
     ELSIF (#statStatus = #STATUS_COMMAND_ABORTED) AND (#statCommandAborted = FALSE) THEN // Commanded functionality has been aborted by another command
       #statDone := FALSE;
       #statBusy := FALSE;
       #statCommandAborted := TRUE;
       #statError := FALSE;
       #diagnostics.stateNumber := #statFBState;
       #diagnostics.status := #statStatus;
       #diagnostics.subfunctionStatus := #statSubfunctionStatus;
       #statFBState := #FB_STATE_NO_PROCESSING; // Switch state machine to "no processing"

       // Reset pointer
       #lineBuffer.pointers.addPointer := 0;
       #lineBuffer.pointers.addPointerRestarted := FALSE;
       #lineBuffer.pointers.bufferLocked := FALSE;
       IF #lineBuffer.info.fileState <> "LKINLANG_FILE_STATE_RUNNING"
         AND #lineBuffer.info.fileState <> "LKINLANG_FILE_STATE_RUNNING_LOADING" THEN
         #lineBuffer.pointers.ignoreAddPointer := TRUE;
       END_IF;

       // Set file state
       #lineBuffer.info.fileState := "LKINLANG_FILE_STATE_STOPPED";


     ELSIF (#statCommandAborted = TRUE) AND (#tempStop = FALSE) THEN
       #statDone := FALSE;
       #statBusy := FALSE;
       #statCommandAborted := FALSE;
       #statError := FALSE;
       #statStatus := #STATUS_NO_CALL;

       // Reset file state
       #lineBuffer.info.fileState := "LKINLANG_FILE_STATE_IDLE";

     ELSIF (#tempExecuteCardToPlc = FALSE) AND (#tempExecutePlcToCard = FALSE) AND ((#statDone = TRUE) OR (#statError = TRUE)) THEN
       #statDone := FALSE;
       #statBusy := FALSE;
       #statCommandAborted := FALSE;
       #statError := FALSE;
       #statStatus := #STATUS_NO_CALL;

       IF #lineBuffer.info.fileState = "LKINLANG_FILE_STATE_STOPPED" THEN
         // Reset file state
         #lineBuffer.info.fileState := "LKINLANG_FILE_STATE_IDLE";
       END_IF;
     END_IF;


     // Write static values to outputs
     #done := #statDone;
     #busy := #statBusy;
     #dataTransferStopped := #statCommandAborted;
     #error := #statError;
     #status := #statStatus;

   END_REGION OUTPUTS

   //--------------------------------------------------------------------
   // End of Block LKinLang_FileHandler
   //--------------------------------------------------------------------
END_FUNCTION_BLOCK

FUNCTION_BLOCK "LKinLang_ProgramLineDisplay"   // FB35452, SCL
TITLE = LKinLang_ProgramLineDisplay
{ S7_Optimized_Access := 'TRUE' }
AUTHOR : tech.team.motioncontrol@siemens.com
FAMILY : LKinLang
VERSION : 1.0
// This FB shows the current parsed, buffered and active line
   VAR_INPUT
      enable : Bool;   // TRUE: Enable functionality of FB
      activeCmdNo : DInt;   // Currently active command number (FB MovePath output)
      movePathStatus : Word;   // Current status output of FB MovePath
   END_VAR
   VAR_OUTPUT
      valid : Bool;   // TRUE: Valid set of output values available at the FB
      busy : Bool;   // TRUE: FB is not finished and new output values can be expected
      error : Bool;   // TRUE: An error occurred during the execution of the FB
      status : Word := 16#7000;   // 16#0000 - 16#7FFF: Status of the FB, 16#8000 - 16#FFFF: Error identification
      parsedLineNo : UDInt;   // Last parsed line number
      parsedLine : String;   // Last parsed line
      bufferedLineNo : UDInt;   // Last buffered line number (internal storage of FB MovePath)
      bufferedLine : String;   // Last buffered line (internal storage of FB MovePath)
      activeLineNo : UDInt;   // Currently active line number
      activeLine : String;   // Currently active line
   END_VAR
   VAR_IN_OUT
      lineBuffer : "LKinLang_typeLineBuffer";   // LineBuffer connection
      pathData : "LKinCtrl_typePathData_advanced";   // PathData connection
   END_VAR
   VAR
      statEnableOld : Bool;   // Old value of 'enable' input for edge detection
      statValid : Bool;   // Static value for output 'valid'
      statBusy : Bool;   // Static value for output 'busy'
      statError : Bool;   // Static value for output 'error'
      statStatus : Word := 16#7000;   // Static value for output 'status'
      statParsedLine : String;   // Static value for output 'parsedLine'
      statParsedLineNo : UDInt;   // Static value for output 'parsedLineNo'
      statBufferedLine : String;   // Static value for output 'bufferedLine'
      statBufferedLineNo : UDInt;   // Static value for output 'bufferedLineNo'
      statActiveLine : String;   // Static value for output 'activeLine'
      statActiveLineNo : UDInt;   // Static value for output 'activeLineNo'
      statErrorUserCleared : Bool;   // Error occurred that can only be solved by user; rising edge at enable input necessary
      statErrorAutoCleared : Bool;   // Error occurred that can be acknowledged by FB
      statFBState : DInt := 0;   // State in the state machine of the FB
      statDisablingCompleted : Bool;   // TRUE: Disabling has been completed
      statAddPointerPathOld : DInt;   // Last value of PathData add pointer
      statRetPointerPathOld : DInt;   // Last value of PathData retrieve pointer
      statActiveCmdNoOld : DInt;   // Last value of active command number
      statRetPointerLineOld : DInt;   // Last value of LineBuffer retrieve pointer
      statBufferIndex : DInt;   // Counter for internal buffer
      statFirstBufferEntry : DInt;   // Static storage for first entry in internal buffer
      statFirstActiveBufferEntry : DInt;   // Static storage for first active entry in internal buffer
      statParsingDone : Bool;   // TRUE: FB Parser is done
      statBufferingDone : Bool;   // TRUE: FB MovePath has copied all commands from PathData
      statMovePathDone : Bool;   // TRUE: FB MovePath has executed all commands from PathData
      statPathDataLines : Array[1.."LKINCTRL_NO_OF_PATHDATA_ELEMENTS_ADVANCED"] of String["LKINLANG_LENGTH_OF_ASCII_LINE_STRING"];   // Stores the corresponding lines from PathData
      statPathDataLineNo : Array[1.."LKINCTRL_NO_OF_PATHDATA_ELEMENTS_ADVANCED"] of UDInt;   // Stores the corresponding line numbers from PathData
      statInternalLines : Array[0..#LAST_INDEX_INTERNAL] of String["LKINLANG_LENGTH_OF_ASCII_LINE_STRING"];   // Stores the corresponding lines from FB MovePath internal buffer
      statInternalLineNo : Array[0..#LAST_INDEX_INTERNAL] of UDInt;   // Stores the corresponding line numbers from FB MovePath internal buffer
   END_VAR
   VAR_TEMP
      tempEnable : Bool;   // Temporary value for input 'enable'
      tempAddPointerPath : DInt;   // Temporary value for input 'PathData.pointers.addPointer'
      tempRetPointerPath : DInt;   // Temporary value for input 'PathData.pointers.retrievePointer'
      tempAddPointerLine : DInt;   // Temporary value for input 'LineBuffer.pointers.addPointer'
      tempRetPointerLine : DInt;   // Temporary value for input 'LineBuffer.pointers.retrievePointer'
      tempActiveCmdNo : DInt;   // Temporary value for input 'activeCmdNo'
      tempMovePathStatus : DWord;   // Temporary value for input 'movePathStatus'
      tempIndex : DInt;   // Temporary counter
   END_VAR
   VAR CONSTANT
      FB_STATE_NO_PROCESSING : DInt := 0;   // FB state: No processing
      FB_STATE_PROCESSING : DInt := 50;   // FB state: Processing
      FB_STATE_DISABLING : DInt := 90;   // FB state: Disabling
      STATUS_NO_CALL : Word := 16#7000;   // No job being currently processed
      STATUS_FIRST_CALL : Word := 16#7001;   // First call after incoming new job (rising edge 'enable')
      STATUS_SUBSEQUENT_CALL : Word := 16#7002;   // Subsequent call during active processing without further details
      ERR_UNDEFINED_STATE : Word := 16#8600;   // Error due to an undefined state in state machine
      LAST_INDEX_INTERNAL : DInt := 19;   // Last index of internal array
   END_VAR
BEGIN
   //=============================================================================
   // SIEMENS AG
   // (c)Copyright 2020
   //-----------------------------------------------------------------------------
   // Library:       LKinLang
   // Tested with:   S7-1517T-3 PN/DP
   // Engineering:   TIA Portal V16
   // Restrictions:  -
   // Requirements:  -
   // Functionality: This FB shows the current parsed, buffered and active line
   //-----------------------------------------------------------------------------
   // Change log table:
   // Version      Date        Expert in charge    Changes applied
   // 01.00.00     03.12.2020  FR                  First created version
   //=============================================================================

   // Work with temporary value / create process image
   #tempEnable := #enable;
   #tempAddPointerPath := #pathData.pointers.addPointer;
   #tempRetPointerPath := #pathData.pointers.retrievePointer;
   #tempAddPointerLine := #lineBuffer.pointers.addPointer;
   #tempRetPointerLine := #lineBuffer.pointers.retrievePointer;
   #tempActiveCmdNo := #activeCmdNo;
   #tempMovePathStatus := #movePathStatus;

   REGION ENABLING/DISABLING
       IF (#tempEnable = TRUE) AND (#statStatus = #STATUS_NO_CALL) THEN // Enable FB
           // First call; initialize FB
           #statValid := TRUE;
           #statBusy := TRUE;
           #statError := FALSE;
           #statErrorUserCleared := FALSE;
           #statErrorAutoCleared := FALSE;
           #statStatus := #STATUS_FIRST_CALL;

           #statFBState := #FB_STATE_PROCESSING; // State machine - start functionality

           // Reset of variables, diagnostics, etc.
           #statDisablingCompleted := FALSE;

           // Reset "old" variables
           #statAddPointerPathOld := 0;
           #statRetPointerPathOld := 0;
           #statActiveCmdNoOld := 0;
           #statRetPointerLineOld := 0;

           // Reset counter / index
           #statBufferIndex := 0;
           #statFirstBufferEntry := 0;
           #statFirstActiveBufferEntry := 0;

           // Reset status bits
           #statParsingDone := FALSE;
           #statBufferingDone := FALSE;

           // Reset arrays
           FOR #tempIndex := 0 TO #LAST_INDEX_INTERNAL DO
               #statInternalLines[#tempIndex] := '';
               #statInternalLineNo[#tempIndex] := 0;
           END_FOR;
           FOR #tempIndex := 1 TO "LKINCTRL_NO_OF_PATHDATA_ELEMENTS_ADVANCED" DO
               #statPathDataLines[#tempIndex] := '';
               #statPathDataLineNo[#tempIndex] := 0;
           END_FOR;

       ELSIF (#tempEnable = FALSE) AND (#statEnableOld = TRUE) THEN // Disable FB 
           #statFBState := #FB_STATE_DISABLING;

       ELSIF (#statStatus = #STATUS_FIRST_CALL) THEN // Set status identifier of subsequent call
           #statStatus := #STATUS_SUBSEQUENT_CALL;
       END_IF;

       // Edge detection 'enable' input
       #statEnableOld := #tempEnable;
   END_REGION ENABLING/DISABLING

   IF (#statStatus = #STATUS_NO_CALL) THEN // Nothing to do -> End here to reduce "system load"
       RETURN;
   END_IF;

   REGION STATE_MACHINE
       CASE #statFBState OF // State machine of FB
           #FB_STATE_NO_PROCESSING: // No processing active (Note: this state must always be present and left empty)
               ;

           #FB_STATE_PROCESSING: // Processing active
               // -----------------------------------------------------------------
               // If a new pathData command was added then store the corresponding
               // lineBuffer entry in the internal pathData buffer
               // 
               // Also check if parsing has finished
               // -----------------------------------------------------------------
               REGION STORE_LINES_INTERNAL
                   // Calculate index
                   IF #tempRetPointerLine > 0 THEN
                       // regular 
                       #tempIndex := #tempRetPointerLine;
                       #statParsingDone := FALSE;
                   ELSIF #tempRetPointerLine = 0 AND #statRetPointerLineOld <> 0 THEN
                       // Parser finished --> retrieve pointer is reset instantly --> Use old value
                       #tempIndex := #statRetPointerLineOld;
                       #statParsingDone := TRUE;
                   ELSE
                       #tempIndex := 0;
                   END_IF;

                   // Check if new pathData command was added
                   IF #tempAddPointerPath <> #statAddPointerPathOld AND #tempAddPointerPath > 0 AND #tempIndex <> 0 THEN
                       // Store the corresponding line in path data line buffer
                       #statPathDataLines[#tempAddPointerPath] := #lineBuffer.lines[#tempIndex].content;
                       #statPathDataLineNo[#tempAddPointerPath] := #lineBuffer.lines[#tempIndex].number;
                   END_IF;

                   // Reset variables if parsing is done
                   IF #statParsingDone THEN
                       ; // Something to reset here?
                   END_IF;
               END_REGION STORE_LINES_INTERNAL


               // -----------------------------------------------------------------
               // Get the currently parsed line information from the lineBuffer
               // -----------------------------------------------------------------
               REGION PARSED_LINE
                   // Check retrieve pointer in lineBuffer --> parsed line 
                   IF #tempRetPointerLine > 0 THEN
                       #statParsedLine := #lineBuffer.lines[#tempRetPointerLine].content;
                       #statParsedLineNo := #lineBuffer.lines[#tempRetPointerLine].number;
                   END_IF;
               END_REGION PARSED_LINE


               // -----------------------------------------------------------------
               // Get the currently buffered line (buffered in MovePath) information from the internal pathData buffer
               // Store the information in the next buffer (statInternalBuffer)
               // --> Buffered lines / cmds in MovePath
               // -----------------------------------------------------------------
               REGION BUFFERED_LINE
                   // Check if buffering was done and set first buffer entry
                   IF #statBufferingDone AND #tempRetPointerPath > 0 THEN
                       #statFirstBufferEntry := #statBufferIndex;
                   END_IF;

                   // Calculate index for pathData lines
                   IF #tempRetPointerPath > 0 AND #statRetPointerPathOld = 0 THEN
                       // First cycle of movePath could process more than one command
                       FOR #tempIndex := 1 TO #tempRetPointerPath DO
                           #statBufferedLine := #statInternalLines[#statBufferIndex] := #statPathDataLines[#tempIndex];
                           #statBufferedLineNo := #statInternalLineNo[#statBufferIndex] := #statPathDataLineNo[#tempIndex];
                           // Count buffer index from 0 to 19
                           #statBufferIndex += 1;
                           #statBufferIndex := #statBufferIndex MOD (#LAST_INDEX_INTERNAL + 1);
                       END_FOR;
                       #tempIndex := 0;
                       #statBufferingDone := FALSE;

                   ELSIF #tempRetPointerPath > 0 AND #statRetPointerPathOld <> #tempRetPointerPath THEN
                       // Regular
                       #tempIndex := #tempRetPointerPath;
                       #statBufferingDone := FALSE;

                   ELSIF #tempRetPointerPath = 0 AND #statRetPointerPathOld <> 0 THEN
                       // MovePath has reached cmdType = -1 --> RetPointerPath is reset in this cycle and does not point to the -1 cmd
                       IF #statRetPointerPathOld + 1 <= "LKINCTRL_NO_OF_PATHDATA_ELEMENTS_ADVANCED" THEN
                           // Regular
                           #tempIndex := #statRetPointerPathOld + 1;
                       ELSE
                           // Old retPointer was last index so the -1 cmd should be on first index
                           #tempIndex := 1;
                       END_IF;
                       // Set buffering done
                       #statBufferingDone := TRUE;
                   ELSE
                       // Both pointer variables are 0 --> Nothing to do
                       #tempIndex := 0;
                   END_IF;

                   // Check retrieve pointer in path data --> buffered line
                   IF #tempIndex <> 0 THEN
                       #statBufferedLine := #statInternalLines[#statBufferIndex] := #statPathDataLines[#tempIndex];
                       #statBufferedLineNo := #statInternalLineNo[#statBufferIndex] := #statPathDataLineNo[#tempIndex];
                       // Count buffer index from 0 to 19
                       #statBufferIndex += 1;
                       #statBufferIndex := #statBufferIndex MOD (#LAST_INDEX_INTERNAL + 1);
                   END_IF;

                   IF #statBufferingDone THEN
                       ; // Something to reset here?
                   END_IF;
               END_REGION BUFFERED_LINE


               // -----------------------------------------------------------------
               // Get the currently active line (active in MovePath) information from the internal buffer
               // -----------------------------------------------------------------
               REGION ACTIVE_LINE
                   // Counting logic
                   (*
                   // activeCmd = 1 | counter = 0
                   // activeCmd = 2 | counter = 1
                   // activeCmd = 3 | counter = 2
                   // activeCmd = 10 | counter = 9
                   // activeCmd = 11 | counter = 10
                   // activeCmd = 19 | counter = 18
                   // activeCmd = 20 | counter = 19
                   // activeCmd = 21 | counter = 0
                   // activeCmd = 22 | counter = 1
                   // activeCmd = 25 | counter = 4
                   // activeCmd = 29 | counter = 8
                   // activeCmd = 30 | counter = 9
                   // activeCmd = 31 | counter = 10
                   // activeCmd = 39 | counter = 18
                   // activeCmd = 40 | counter = 19
                   // activeCmd = 41 | counter = 0
                   *)

                   // Check if movePath is done
                   IF #tempMovePathStatus = 16#0000 OR #tempMovePathStatus = 16#7000 THEN
                       #statMovePathDone := TRUE;
                   END_IF;

                   // If active cmd changes, reset movePath done
                   IF #tempActiveCmdNo <> #statActiveCmdNoOld THEN
                       #statMovePathDone := FALSE;
                   END_IF;

                   // If active cmd is less then last active cmd then update first buffer entry
                   IF #tempActiveCmdNo < #statActiveCmdNoOld THEN
                       #statFirstActiveBufferEntry := #statFirstBufferEntry;
                   END_IF;

                   // Active line
                   IF #tempActiveCmdNo > 0 THEN
                       // tempIndex shall run from 0 to 19
                       #tempIndex := (#statFirstActiveBufferEntry + #tempActiveCmdNo - 1) MOD (#LAST_INDEX_INTERNAL + 1);
                       // MovePath is done
                       IF #statMovePathDone = TRUE THEN
                           IF #tempIndex < #LAST_INDEX_INTERNAL THEN
                               #tempIndex += 1;
                           ELSE
                               #tempIndex := 1;
                           END_IF;
                       END_IF;
                       #statActiveLine := #statInternalLines[#tempIndex];
                       #statActiveLineNo := #statInternalLineNo[#tempIndex];
                   END_IF;
               END_REGION ACTIVE_LINE


           #FB_STATE_DISABLING: // Disabling active
               // TODO: Disabling, e.g. closing connections, etc.
               // When disabling is complete the bit #statDisablingCompleted must be set
               #statDisablingCompleted := TRUE;

           ELSE // Undefined state in state machine reached
               #statStatus := #ERR_UNDEFINED_STATE;
               #statErrorUserCleared := TRUE;
       END_CASE;
   END_REGION STATE_MACHINE

   REGION STORE_OLD
       // Store old
       #statAddPointerPathOld := #tempAddPointerPath;
       #statRetPointerPathOld := #tempRetPointerPath;
       #statRetPointerLineOld := #tempRetPointerLine;
       #statActiveCmdNoOld := #tempActiveCmdNo;
   END_REGION STORE_OLD

   REGION OUTPUTS
       // Write outputs
       IF (#statDisablingCompleted = TRUE) THEN
           // Reset outputs if disabling completed
           #statValid := FALSE;
           #statBusy := FALSE;
           #statError := FALSE;
           #statErrorUserCleared := FALSE;
           #statErrorAutoCleared := FALSE;
           #statStatus := #STATUS_NO_CALL;
           // Reset application specific outputs
           #statParsedLine := #statBufferedLine := #statActiveLine := '';
           #statParsedLineNo := #statBufferedLineNo := #statActiveLineNo := 0;

       ELSIF (#statErrorUserCleared = TRUE) AND (#statError = FALSE) THEN
           // Error can only be cleared by user; rising edge at enable input is needed to continue 
           #statValid := FALSE;
           #statBusy := FALSE;
           #statError := TRUE;
           #statFBState := #FB_STATE_NO_PROCESSING; // Switch state machine to "no processing"

       ELSIF (#statErrorAutoCleared = TRUE) AND (#statError = FALSE) THEN
           // Error can be reset by FB automatically  
           #statValid := FALSE;
           #statBusy := TRUE;
           #statError := TRUE;
           // TODO: Handling of autocleared error

       ELSIF (#statErrorAutoCleared = FALSE) AND (#statErrorUserCleared = FALSE) AND (#statError = TRUE) THEN
           // If autocleared error is acknowledged
           #statValid := TRUE;
           #statBusy := TRUE;
           #statError := FALSE;
           #statStatus := #STATUS_SUBSEQUENT_CALL;
       END_IF;

       // Write static values to outputs
       #valid := #statValid;
       #busy := #statBusy;
       #error := #statError;
       #status := #statStatus;
       // Write application specific static values to outputs
       #parsedLine := #statParsedLine;
       #parsedLineNo := #statParsedLineNo;
       #bufferedLine := #statBufferedLine;
       #bufferedLineNo := #statBufferedLineNo;
       #activeLine := #statActiveLine;
       #activeLineNo := #statActiveLineNo;
   END_REGION OUTPUTS
END_FUNCTION_BLOCK

// folder: LKinLang_Blocks/LKinLang_LanguageDefinition

FUNCTION "LKinLang_SelectLangPackage" : Void   // FC35450, SCL
TITLE = LKinLang_SelectLangPackage
{ S7_Optimized_Access := 'TRUE' }
AUTHOR : tech.team.motioncontrol@siemens.com
FAMILY : LKinLang
VERSION : 1.1
// The FC selects a language package and definition of user parameters and returns the languages
// syntax by parameter definition, separators, mergers and valid counts
   VAR_INPUT
      language : Int;   // Selected Language
   END_VAR
   VAR_OUTPUT
      separators : Array[1.."LKINLANG_NUMBER_OF_SEPARATORS"] of Byte;   // Found separators
      mergers : Array[1.."LKINLANG_NUMBER_OF_MERGERS"] of Byte;   // Found mergers
      validCounts : "LKinLang_typePathDataElementCounter";   // Array which defines how often a parameter can be set
      variableDeclarations : "LKinLang_typeVariableDeclaration";   // Syntax how to declare local variables
      keyToken : "LKinLang_typeKeyToken";   // Keywords for different commands
   END_VAR
   VAR_IN_OUT
      parameterDefinition : "LKinLang_typeParameterDefinition";   // Found command definition
      parameterNumber : Int;   // Parameter number
      parameterDefaults : Variant;   // Parameter defaults
   END_VAR
   VAR_TEMP
      tempConditionCounter : Int;   // Temprary counter
      tempGCodeDefaults : REF_TO "LKinLang_typeGCodeDefaults";   // Reference to GCode defaults
      tempUserDefinedDefaults : REF_TO "LKinLang_typeUserDefinedDefaults";   // Reference to UserDefined defaults
   END_VAR
   VAR CONSTANT
      ERR_WRONG_DEFAULTS : Int := -998;   // Error due to missing or wrong default connection
      ERR_LANG_NOT_DEFINED : Int := -999;   // Error selected language not defined
      FIRST_USERDEF_GCODE : DInt := 1;   // First parameter number for user defined GCode
      LAST_USERDEF_GCODE : DInt := 99;   // Last parameter number for user defined GCode
      FIRST_PREDEF_GCODE : DInt := 100;   // First parameter number for PreDefined GCode
      LAST_PREDEF_GCODE : DInt := 199;   // Last parameter number for PreDefined GCode
      FIRST_USERDEF_LANG : DInt := 1;   // First parameter number for user defined language
      LAST_USERDEF_LANG : DInt := 199;   // Last parameter number for user defined language
      END_OF_CASE : DInt := 200;   // End of case
   END_VAR
BEGIN
   //==========================================================================================
   // SIEMENS AG
   // (c)Copyright 2020 All Rights Reserved
   //------------------------------------------------------------------------------------------
   // Library: LKinLang
   // Tested with: S7-1517T-3 PN/DP
   // Engineering: TIA Portal V15
   // Restrictions: ---
   // Requirements: S7-1500T FW 2.5
   // Functionality: LKinLang_SelecLangPackage
   // The FC selects a language package and definition of user parameters and returns the languages
   // syntax by parameter definition, separators, mergers and valid counts
   // 
   // Support: tech.team.motioncontrol@siemens.com
   // Note: Parameter comments are only available in language 'English (United States)'
   //------------------------------------------------------------------------------------------
   // Change log table:
   // Version    Date          Expert in charge    Changes applied
   // 01.00.00   28.05.2019    FR                  First created version
   // 01.00.02   29.07.2019    FR                  Removed empty path data element from interface; parameter definition now InOut
   // 01.00.03   19.03.2020    FR                  Added valueFlagsCount to UserDefined
   // 01.01.00   24.03.2020    FR                  Added variableDeclaration and KeyToken
   // 01.02.00   02.11.2020    FR                  Added IF,FOR,WHILE,SUB to KeyToken
   //===========================================================================================

   // Select language package with Parser input "language"
   // 
   CASE #language OF
     "LKINLANG_LANGPACK_GCODE":  // G-Code language package
       REGION GCODE_LANGUAGE

         // Check type of variant input
         IF TypeOf(#parameterDefaults) = LKinLang_typeGCodeDefaults THEN
           #tempGCodeDefaults ?= #parameterDefaults;
         ELSE
           // Error wrong data type
           #parameterNumber := #ERR_WRONG_DEFAULTS;
           RETURN;
         END_IF;

         REGION SEPARATORS_MERGERS
           // Separators
           #separators[1] := 16#20; // Space
           #separators[2] := 16#26; // &
           #separators[3] := 16#3D; // =
           #separators[4] := 16#3E; // >
           #separators[5] := 16#3C; // <
           #separators[6] := 16#28; // (
           #separators[7] := 16#29; // )
           #separators[8] := 16#2F; // /
           #separators[9] := 16#2A; // *
           #separators[10] := 16#2B; // +
           #separators[11] := 16#2D; // -
           #separators[12] := 16#7C; // |
           #separators[13] := 16#3A; // :
           #separators[14] := 16#5E; // ^
           #separators[15] := 16#2C; // ,

           // Mergers (to enable e.g. Test_1)
           #mergers[1] := 16#5F; // _

         END_REGION SEPARATORS_MERGERS

         REGION KEY_TOKEN
           // Define keyword token
           // Define local variable data type token --> Used below as "_type_"
           #keyToken.tokenBool := 'BOOL';
           #keyToken.tokenDInt := 'DINT';
           #keyToken.tokenLReal := 'LREAL';

           // Define keyword for using interface variables
           #keyToken.tokenInterfaceVarBool := '%B';
           #keyToken.tokenInterfaceVarDInt := '%DI';
           #keyToken.tokenInterfaceVarLReal := '%LR';

           // Keywords for jumps, label(jump target) and stopre (sync movePath and Parser)
           #keyToken.tokenJump := 'GOTO';
           #keyToken.tokenJumpConditional := 'GOTOC';
           #keyToken.tokenJumpTarget := 'LABEL';
           #keyToken.tokenPreprocessingStop := 'STOPRE';

           // Keywords loops, jumps, subprogram
           #keyToken.tokenIf := 'IF';
           #keyToken.tokenEndIf := 'ENDIF';
           #keyToken.tokenWhile := 'WHILE';
           #keyToken.tokenEndWhile := 'ENDWHILE';
           #keyToken.tokenFor := 'FOR';
           #keyToken.tokenQuantity := 'TO';
           #keyToken.tokenIncrement := 'STEP';
           #keyToken.tokenEndFor := 'ENDFOR';
           #keyToken.tokenStartSub := 'SUB';
           #keyToken.tokenEndSub := 'ENDSUB';
           #keyToken.tokenCallSub := 'CALL';
           #keyToken.tokenReturnSub := 'RETURN';
         END_REGION KEY_TOKEN

         REGION VARIABLE_DEFINITION
           // Local variable declaration
           // Use _name_ to specify the position of the variable name
           // Use _type_ to specify the position of the variable data type
           // Possible data types:
           // - BOOL
           // - DINT
           // - LREAL

           #variableDeclarations.localVariables := 'DEF _type_ _name_';
           #variableDeclarations.globalVariables := 'DEF GLOBAL _type_ _name_';
         END_REGION VARIABLE_DEFINITION


         REGION VALID_COUNTS
           #validCounts.cmdType := 1; // One change of cmdType allowed per PathData command
           #validCounts.cmdName := 1;

           #validCounts.cmdCoordinates.cartesianPosition.x := 1;
           #validCounts.cmdCoordinates.cartesianPosition.y := 1;
           #validCounts.cmdCoordinates.cartesianPosition.z := 1;
           #validCounts.cmdCoordinates.cartesianPosition.a := 1;
           #validCounts.cmdCoordinates.coordSystem := 1;

           #validCounts.cmdParameters.bufferMode := 1;
           #validCounts.cmdParameters.dynamicAdaption := 1;
           #validCounts.cmdParameters.orientationDirection := 1;

           #validCounts.cmdParameters.offsetParameters.mainPathPlane := 1;
           #validCounts.cmdParameters.offsetParameters.offsetParaNo := 1;

           #validCounts.cmdParameters.pathDynamics.velocity := 1;
           #validCounts.cmdParameters.pathDynamics.acceleration := 1;
           #validCounts.cmdParameters.pathDynamics.deceleration := 1;
           #validCounts.cmdParameters.pathDynamics.jerk := 1;

           #validCounts.cmdParameters.circleParameters.arc := 1;
           #validCounts.cmdParameters.circleParameters.circlePlane := 1;
           #validCounts.cmdParameters.circleParameters.circMode := 1;
           #validCounts.cmdParameters.circleParameters.auxPoint[1] := 1;
           #validCounts.cmdParameters.circleParameters.auxPoint[2] := 1;
           #validCounts.cmdParameters.circleParameters.auxPoint[3] := 1;
           #validCounts.cmdParameters.circleParameters.pathChoice := 1;
           #validCounts.cmdParameters.circleParameters.radius := 1;

           #validCounts.cmdParameters.transitionParameters[1] := 1;
           #validCounts.cmdParameters.transitionParameters[2] := 1;
           #validCounts.cmdParameters.transitionParameters[3] := 1;
           #validCounts.cmdParameters.transitionParameters[4] := 1;
           #validCounts.cmdParameters.transitionParameters[5] := 1;

           #validCounts.setFlags.flag := "LKINCTRL_NO_OF_CMD_SETFLAGS";
           #validCounts.setFlags.flagMode := "LKINCTRL_NO_OF_CMD_SETFLAGS";
           #validCounts.setFlags.remainingDistance := "LKINCTRL_NO_OF_CMD_SETFLAGS";

           #validCounts.valueFlags.flag := "LKINCTRL_NO_OF_CMD_VALUEFLAGS";
           #validCounts.valueFlags.value := "LKINCTRL_NO_OF_CMD_VALUEFLAGS";
           #validCounts.valueFlags.flagMode := "LKINCTRL_NO_OF_CMD_VALUEFLAGS";
           #validCounts.valueFlags.remainingDistance := "LKINCTRL_NO_OF_CMD_VALUEFLAGS";
         END_REGION VALID_COUNTS


         REGION PARAMETER_DEFINITION
           // Definiton:
           // Case of ParameterNo = -1 --> End of Case
           // Case of ParameterNo = -2 --> Missing Definition (Else branch)
           // 
           //
           //                                   31   27   23   19   15   11   7    3
           // Properties                        |    |    |    |    |    |    |    |
           // tempCmdDefinition.properties := 2#0000_0000_0000_0000_0000_0000_0000_0000;
           // List of properties:
           // X0: 0=Config CMD, 1=Motion CMD
           // X1: 1=CMD Modal
           // X2: 1=PRG Modal
           // X3: 1=Check limits
           // 
           // X4: 1=Equation allowed
           // X5: 1=Switch to Absolute Position
           // X6: 1=Switch to Relative Positions
           // X7: reserved

           CASE #parameterNumber OF
             #FIRST_USERDEF_GCODE..#LAST_USERDEF_GCODE: // User defined GCode
               REGION USER_DEFINED_GCODE
                 "LKinLang_UserDefinedGCode"(parameterNo := #parameterNumber,
                                             parameterDefinition := #parameterDefinition,
                                             parameterDefaults := #tempGCodeDefaults<?OpDeref?>);
               END_REGION USER_DEFINED_GCODE

             #FIRST_PREDEF_GCODE..#LAST_PREDEF_GCODE: // PreDefined GCode
               REGION PRE_DEFINED_GCODE
                 "LKinLang_LangPackageGCode"(parameterDefinition := #parameterDefinition,
                                             parameterNo := #parameterNumber,
                                             parameterDefaults := #tempGCodeDefaults<?OpDeref?>);
               END_REGION PRE_DEFINDED_GCODE

             #END_OF_CASE: // 200
               // End 0f parameter definition reached
               #parameterNumber := -1; // abort searching

             ELSE  // Statement section ELSE
               // invalid case number
               #parameterNumber := -2;
           END_CASE;
         END_REGION PARAMETER_DEFINITION

         // ---------------------------------------------------
         // End of GCode
         // ---------------------------------------------------
       END_REGION GCODE_LANGUAGE

     "LKINLANG_LANGPACK_USER": // User defined language (completely user defined)
       REGION USER_DEFINED_LANGUAGE

         // Check type of variant input
         IF TypeOf(#parameterDefaults) = LKinLang_typeUserDefinedDefaults THEN
           #tempUserDefinedDefaults ?= #parameterDefaults;
         ELSE
           ; // Error wrong data type
           #parameterNumber := #ERR_WRONG_DEFAULTS;
           RETURN;
         END_IF;

         REGION SEPARATORS_MERGERS
           // Separators
           #separators[1] := 16#20; // Space
           #separators[2] := 16#26; // &
           #separators[3] := 16#3D; // =
           #separators[4] := 16#3E; // >
           #separators[5] := 16#3C; // <
           #separators[6] := 16#28; // (
           #separators[7] := 16#29; // )
           #separators[8] := 16#2F; // /
           #separators[9] := 16#2A; // *
           #separators[10] := 16#2B; // +
           #separators[11] := 16#2D; // -
           #separators[12] := 16#7C; // |
           #separators[13] := 16#3A; // :
           #separators[14] := 16#5E; // ^
           #separators[15] := 16#2C; // ,

           // Mergers (to enable e.g. Test_1)
           #mergers[1] := 16#5F; // _
         END_REGION SEPARATORS_MERGERS

         REGION KEY_TOKEN
           // Define keyword token
           // Define local variable data type token --> Used below as "_type_"
           #keyToken.tokenBool := 'BOOL';
           #keyToken.tokenDInt := 'DINT';
           #keyToken.tokenLReal := 'LREAL';

           // Define keyword for using interface variables
           #keyToken.tokenInterfaceVarBool := '%B';
           #keyToken.tokenInterfaceVarDInt := '%DI';
           #keyToken.tokenInterfaceVarLReal := '%LR';

           // Keywords for jumps, label(jump target) and stopre (sync movePath and Parser)
           #keyToken.tokenJump := 'GOTO';
           #keyToken.tokenJumpConditional := 'GOTOC';
           #keyToken.tokenJumpTarget := 'LABEL';
           #keyToken.tokenPreprocessingStop := 'STOPRE';

           // Keywords loops, jumps, subprogram
           #keyToken.tokenIf := 'IF';
           #keyToken.tokenEndIf := 'ENDIF';
           #keyToken.tokenWhile := 'WHILE';
           #keyToken.tokenEndWhile := 'ENDWHILE';
           #keyToken.tokenFor := 'FOR';
           #keyToken.tokenQuantity := 'TO';
           #keyToken.tokenIncrement := 'STEP';
           #keyToken.tokenEndFor := 'ENDFOR';
           #keyToken.tokenStartSub := 'SUB';
           #keyToken.tokenEndSub := 'ENDSUB';
           #keyToken.tokenCallSub := 'CALL';
           #keyToken.tokenReturnSub := 'RETURN';
         END_REGION KEY_TOKEN

         REGION VARIABLE_DEFINITION
           // Local variable declaration
           // Use _name_ to specify the position of the variable name
           // Use _type_ to specify the position of the variable data type
           // Possible data types:
           // - BOOL
           // - DINT
           // - LREAL

           #variableDeclarations.localVariables := 'DEF _type_ _name_';
           #variableDeclarations.globalVariables := 'DEF GLOBAL _type_ _name_';
         END_REGION VARIABLE_DEFINITION

         REGION VALID_COUNTS
           #validCounts.cmdType := 1; // One change of cmdType allowed per PathData command
           #validCounts.cmdName := 1;

           #validCounts.cmdCoordinates.cartesianPosition.x := 1;
           #validCounts.cmdCoordinates.cartesianPosition.y := 1;
           #validCounts.cmdCoordinates.cartesianPosition.z := 1;
           #validCounts.cmdCoordinates.cartesianPosition.a := 1;
           #validCounts.cmdCoordinates.coordSystem := 1;

           #validCounts.cmdParameters.bufferMode := 1;
           #validCounts.cmdParameters.dynamicAdaption := 1;
           #validCounts.cmdParameters.orientationDirection := 1;

           #validCounts.cmdParameters.offsetParameters.mainPathPlane := 1;
           #validCounts.cmdParameters.offsetParameters.offsetParaNo := 1;

           #validCounts.cmdParameters.pathDynamics.velocity := 1;
           #validCounts.cmdParameters.pathDynamics.acceleration := 1;
           #validCounts.cmdParameters.pathDynamics.deceleration := 1;
           #validCounts.cmdParameters.pathDynamics.jerk := 1;

           #validCounts.cmdParameters.circleParameters.arc := 1;
           #validCounts.cmdParameters.circleParameters.circlePlane := 1;
           #validCounts.cmdParameters.circleParameters.circMode := 1;
           #validCounts.cmdParameters.circleParameters.auxPoint[1] := 1;
           #validCounts.cmdParameters.circleParameters.auxPoint[2] := 1;
           #validCounts.cmdParameters.circleParameters.auxPoint[3] := 1;
           #validCounts.cmdParameters.circleParameters.pathChoice := 1;
           #validCounts.cmdParameters.circleParameters.radius := 1;

           #validCounts.cmdParameters.transitionParameters[1] := 1;
           #validCounts.cmdParameters.transitionParameters[2] := 1;
           #validCounts.cmdParameters.transitionParameters[3] := 1;
           #validCounts.cmdParameters.transitionParameters[4] := 1;
           #validCounts.cmdParameters.transitionParameters[5] := 1;

           #validCounts.setFlags.flag := "LKINCTRL_NO_OF_CMD_SETFLAGS";
           #validCounts.setFlags.flagMode := "LKINCTRL_NO_OF_CMD_SETFLAGS";
           #validCounts.setFlags.remainingDistance := "LKINCTRL_NO_OF_CMD_SETFLAGS";

           #validCounts.valueFlags.flag := "LKINCTRL_NO_OF_CMD_VALUEFLAGS";
           #validCounts.valueFlags.value := "LKINCTRL_NO_OF_CMD_VALUEFLAGS";
           #validCounts.valueFlags.flagMode := "LKINCTRL_NO_OF_CMD_VALUEFLAGS";
           #validCounts.valueFlags.remainingDistance := "LKINCTRL_NO_OF_CMD_VALUEFLAGS";
         END_REGION VALID_COUNTS

         REGION PARAMETER_DEFINITION
           // Definiton:
           // Case of ParameterNo = -1 --> End of Case
           // Case of ParameterNo = -2 --> Missing Definition (Else branch)
           // 
           //
           //                                   31   27   23   19   15   11   7    3
           // Properties                        |    |    |    |    |    |    |    |
           // tempCmdDefinition.properties := 2#0000_0000_0000_0000_0000_0000_0000_0000;
           // List of properties:
           // X0: 0=Config CMD, 1=Motion CMD
           // X1: 1=CMD Modal
           // X2: 1=PRG Modal
           // X3: 1=Check limits
           // 
           // X4: 1=Equation allowed
           // X5: 1=Switch to Absolute Position
           // X6: 1=Switch to Relative Positions
           // X7: reserved


           // Initialize temp variables
           //#tempParameterDefinition.directValues := #pathDataElementEmpty;

           CASE #parameterNumber OF
             #FIRST_USERDEF_LANG..#LAST_USERDEF_LANG: // User defined parameters
               "LKinLang_LangPackageUser"(parameterNo:=#parameterNumber,
                                          parameterDefinition:=#parameterDefinition,
                                          parameterDefaults:=#tempUserDefinedDefaults<?OpDeref?>);

             #END_OF_CASE: // 200
               // End 0f parameter definition reached
               #parameterNumber := -1; // abort searching

             ELSE  // Statement section ELSE
               // invalid case number
               #parameterNumber := -2;
           END_CASE;
         END_REGION PARAMETER_DEFINITION

         // ---------------------------------------------------
         // End of UserDefined language
         // ---------------------------------------------------
       END_REGION USER_DEFINED_LANGUAGE

     ELSE  // Else --> Error language definition missing 
       #parameterNumber := #ERR_LANG_NOT_DEFINED;
   END_CASE;
END_FUNCTION

// folder: LKinLang_Blocks/LKinLang_LanguageDefinition/LKinLang_LangPackGCode

FUNCTION "LKinLang_LangPackageGCode" : Void   // FC35451, SCL
TITLE = LKinLang_LangPackageGCode
{ S7_Optimized_Access := 'TRUE' }
AUTHOR : tech.team.motioncontrol@siemens.com
FAMILY : LKinLang
VERSION : 1.1
// Language definition package containing GCode
   VAR_IN_OUT
      parameterNo : Int;   // Parameter number
      parameterDefinition : "LKinLang_typeParameterDefinition";   // Found parameter definition
      parameterDefaults : "LKinLang_typeGCodeDefaults";   // Parameter defaults
   END_VAR
   VAR_TEMP
      tempConditionCounter : Int;   // Temporary counter variable
   END_VAR
   VAR CONSTANT
      G0 : DInt := 100;   // Fast Lin
      G1 : DInt := 101;   // Lin
      G2 : DInt := 102;   // Circ CW
      G3 : DInt := 103;   // Circ CCW
      G5 : DInt := 105;   // Circ 3D
      G4 : DInt := 104;   // WaitTime
      P : DInt := 110;   // Period for WaitTime
      G17 : DInt := 120;   // XY Plane
      G18 : DInt := 121;   // ZX Plane
      G19 : DInt := 122;   // YZ Plane
      G640 : DInt := 130;   // Geometry blending off
      G641 : DInt := 131;   // Geometry blending with high velocity
      G642 : DInt := 132;   // Geometry blending with low velocity
      G90 : DInt := 150;   // Absolute Position
      G91 : DInt := 151;   // Relativ Position
      G54 : DInt := 152;   // Select OCS1
      G55 : DInt := 153;   // Select OCS2
      G56 : DInt := 154;   // Select OCS3
      G500 : DInt := 155;   // Select WCS
      T : DInt := 160;   // Tool selection
      G40 : DInt := 161;   // Tool off
      G41 : DInt := 162;   // Tool left
      G42 : DInt := 163;   // Tool right
      X : DInt := 170;   // X pos
      Y : DInt := 171;   // Y pos
      Z : DInt := 172;   // Z pos
      "A" : DInt := 173;   // Orientation
      F : DInt := 174;   // Velocity
      ACC : DInt := 175;   // Acceleration
      DEC : DInt := 176;   // Deceleration
      JERK : DInt := 177;   // Jerk
      CR : DInt := 178;   // Circle Radius
      I : DInt := 179;   // Circ Point
      J : DInt := 180;   // Circ Point
      K : DInt := 181;   // Circ Point
      AR : DInt := 182;   // Arc
      BR : DInt := 183;   // Transition Parameter
      "M" : DInt := 190;   // Flag
      H : DInt := 191;   // Value Flag
      M30 : DInt := 199;   // End of PRG
   END_VAR
BEGIN
   //==========================================================================================
   // SIEMENS AG
   // (c)Copyright 2019 All Rights Reserved
   //------------------------------------------------------------------------------------------
   // Library: LKinLang
   // Tested with: S7-1517T-3 PN/DP
   // Engineering: TIA Portal V15
   // Restrictions: ---
   // Requirements: S7-1500T FW 2.5
   // Functionality: LKinLang_LangPackageKinematics
   // Language definition package for kinematics language GCode
   // 
   // Support: tech.team.motioncontrol@siemens.com
   // Note: Parameter comments are only available in language 'English (United States)'
   //------------------------------------------------------------------------------------------
   // Change log table:
   // Version    Date          Expert in charge    Changes applied
   // 01.00.00   28.05.2019    FR                  First created version
   //===========================================================================================
   //
   //  Group Parameter 
   //  10:   F
   //        
   //  20:   G17
   //        G18
   //        G19
   //        
   //  30:   F
   //        P
   //        
   //  40:   T
   //
   //  50:   BR
   //  
   //  60:   I
   //        J
   //        K
   //
   //  70:   X
   //        Y
   //        Z


   CASE #parameterNo OF
       // Motion Parameters (100 - 169)
       // ===========================================================
     #G0: // Rapid Linear
       // Command name definition
       #parameterDefinition.parameterNameString := 'G';
       #parameterDefinition.parameterNameNumber := 0;

       // Properties
       #parameterDefinition.properties := "LKINLANG_MOTION_CMD" + "LKINLANG_CMD_MODAL";
       #parameterDefinition.validCountPerLine := 1;

       // Priorities
       #parameterDefinition.priorities.cmdType := "LKINLANG_PRIO_DEFINED";
       #parameterDefinition.priorities.cmdParameters.pathDynamics.velocity := "LKINLANG_PRIO_CONSTANT";

       // Matching to PathData
       #parameterDefinition.directValues.cmdType := 1;
       #parameterDefinition.directValues.cmdParameters.pathDynamics.velocity := #parameterDefaults.velocityRapidLinear;

     #G1:  // Linear
       // Command name definition
       #parameterDefinition.parameterNameString := 'G';
       #parameterDefinition.parameterNameNumber := 1;

       // Properties
       #parameterDefinition.properties := "LKINLANG_MOTION_CMD" + "LKINLANG_CMD_MODAL";
       #parameterDefinition.validCountPerLine := 1;

       // Conditions
       #tempConditionCounter := 1;
       #parameterDefinition.conditions[#tempConditionCounter].ParameterNumber := #F;
       #parameterDefinition.conditions[#tempConditionCounter].Group := 10;
       #parameterDefinition.conditions[#tempConditionCounter].Mode := "LKINLANG_CONDITION_IN_PROGRAM"; // In program

       // Priorities
       #parameterDefinition.priorities.cmdType := "LKINLANG_PRIO_DEFINED";

       // Matching to PathData
       #parameterDefinition.directValues.cmdType := 1;


     #G2:  // Circ CW --> CircMode 1/2/3
       // Command name definition
       #parameterDefinition.parameterNameString := 'G';
       #parameterDefinition.parameterNameNumber := 2;

       // Properties
       #parameterDefinition.properties := "LKINLANG_MOTION_CMD" + "LKINLANG_CMD_MODAL";
       #parameterDefinition.validCountPerLine := 1;

       // Conditions
       #tempConditionCounter := 1;
       #parameterDefinition.conditions[#tempConditionCounter].ParameterNumber := #G17;
       #parameterDefinition.conditions[#tempConditionCounter].Group := 20;
       #parameterDefinition.conditions[#tempConditionCounter].Mode := "LKINLANG_CONDITION_IN_PROGRAM"; // In program
       #tempConditionCounter += 1;
       #parameterDefinition.conditions[#tempConditionCounter].ParameterNumber := #G18;
       #parameterDefinition.conditions[#tempConditionCounter].Group := 20;
       #parameterDefinition.conditions[#tempConditionCounter].Mode := "LKINLANG_CONDITION_IN_PROGRAM"; // In program
       #tempConditionCounter += 1;
       #parameterDefinition.conditions[#tempConditionCounter].ParameterNumber := #G19;
       #parameterDefinition.conditions[#tempConditionCounter].Group := 20;
       #parameterDefinition.conditions[#tempConditionCounter].Mode := "LKINLANG_CONDITION_IN_PROGRAM"; // In program
       #tempConditionCounter += 1;
       #parameterDefinition.conditions[#tempConditionCounter].ParameterNumber := #F;
       #parameterDefinition.conditions[#tempConditionCounter].Group := 10;
       #parameterDefinition.conditions[#tempConditionCounter].Mode := "LKINLANG_CONDITION_IN_PROGRAM"; // In program


       // Priorities
       // PathChoice and CmdType are defined
       #parameterDefinition.priorities.cmdType := "LKINLANG_PRIO_DEFINED";
       #parameterDefinition.priorities.cmdParameters.circleParameters.pathChoice := "LKINLANG_PRIO_DEFINED";

       // CircMode and circPlane can be changed (G17,G18,G19 / AR,CR,I,J,K)
       #parameterDefinition.priorities.cmdParameters.circleParameters.circlePlane := "LKINLANG_PRIO_DEFAULT";
       #parameterDefinition.priorities.cmdParameters.circleParameters.circMode := "LKINLANG_PRIO_DEFAULT";

